// TIA Portal project "1215C_BREAKOUT_BOARD" (V19)

(* hardware
DEVICE "S7-1200 station_1"  S7-1200 Station
   slot 0: "Rack_0"  S7-1200 Rack  Rack  V1.0
   slot 1: "BREAKOUT_BOARD_PLC"  CPU 1215C DC/DC/DC  6ES7 215-1AG40-0XB0  V4.6
DEVICE "BREAKOUT_BOARD_HMI"  KTP400 Basic PN
   slot 0: "BREAKOUT_BOARD_HMI"  KTP400 Basic PN  6AV2 123-2DB03-0AX0  16.0.0.0
   slot 1: "HMI_RT_1"  KTP400 Basic PN  6AV2 123-2DB03-0AX0  16.0.0.0
   slot 5: "BREAKOUT_BOARD_HMI.IE_CP_1"  PROFINET Interface  16.0.0.0
      slot 1: "PROFINET Interface"  PROFINET Interface
         slot 1: "Port_1"  Port
*)

// ===== PLC "BREAKOUT_BOARD_PLC"  CPU 1215C DC/DC/DC =====

VAR_GLOBAL   // PLC tag table "PLC_Outputs"
   "DQ0.0" AT %Q0.0 : Bool;   // Digital Output
   "DQ0.1" AT %Q0.1 : Bool;   // Digital Output
   "DQ0.2" AT %Q0.2 : Bool;   // Digital Output
   "DQ0.3" AT %Q0.3 : Bool;   // Digital Output
   "DQ0.4" AT %Q0.4 : Bool;   // Digital Output
   "DQ0.5" AT %Q0.5 : Bool;   // Digital Output
   "DQ0.6" AT %Q0.6 : Bool;   // Digital Output
   "DQ0.7" AT %Q0.7 : Bool;   // Digital Output
   "DQ1.0" AT %Q1.0 : Bool;   // Digital Output
   "DQ1.1" AT %Q1.1 : Bool;   // Digital Output
   "AQ0.0" AT %QW64 : Word;   // Analog Output
   "AQ0.1" AT %QW66 : Word;   // Analog Output
END_VAR

VAR_GLOBAL   // PLC tag table "PLC_Inputs"
   "DI0.0" AT %I0.0 : Bool;   // Digital Input
   "DI0.1" AT %I0.1 : Bool;   // Digital Input
   "DI0.2" AT %I0.2 : Bool;   // Digital Input
   "DI0.3" AT %I0.3 : Bool;   // Digital Input
   "DI0.4" AT %I0.4 : Bool;   // Digital Input
   "DI0.5" AT %I0.5 : Bool;   // Digital Input
   "DI0.6" AT %I0.6 : Bool;   // Digital Input
   "DI0.7" AT %I0.7 : Bool;   // Digital Input
   "DI1.0" AT %I1.0 : Bool;   // Digital Input
   "DI1.1" AT %I1.1 : Bool;   // Digital Input
   "DI1.2" AT %I1.2 : Bool;   // Digital Input
   "DI1.3" AT %I1.3 : Bool;   // Digital Input
   "DI1.4" AT %I1.4 : Bool;   // Digital Input
   "DI1.5" AT %I1.5 : Bool;   // Digital Input
   "AI0.0" AT %IW64 : Word;   // Analog Input
   "AI0.1" AT %IW66 : Word;   // Analog Input
END_VAR

VAR_GLOBAL   // PLC tag table "System_Tags"
   "Clock_Byte" AT %MB0 : Byte;
   "Clock_10Hz" AT %M0.0 : Bool;
   "Clock_5Hz" AT %M0.1 : Bool;
   "Clock_2.5Hz" AT %M0.2 : Bool;
   "Clock_2Hz" AT %M0.3 : Bool;
   "Clock_1.25Hz" AT %M0.4 : Bool;
   "Clock_1Hz" AT %M0.5 : Bool;
   "Clock_0.625Hz" AT %M0.6 : Bool;
   "Clock_0.5Hz" AT %M0.7 : Bool;
   "System_Byte" AT %MB1 : Byte;
   "FirstScan" AT %M1.0 : Bool;
   "DiagStatusUpdate" AT %M1.1 : Bool;
   "AlwaysTRUE" AT %M1.2 : Bool;
   "AlwaysFALSE" AT %M1.3 : Bool;
END_VAR

VAR_GLOBAL   // PLC tag table "Trigger_Tags"
   "xAQ_Trig" AT %M2.0 : Bool;
   "xTrig2" AT %M2.1 : Bool;
   "xTrig3" AT %M2.2 : Bool;
   "xTrig4" AT %M2.3 : Bool;
   "xTrig5" AT %M2.4 : Bool;
END_VAR

// folder: WS01_TVET_Workstation/00-I/O_Mapping

DATA_BLOCK "DB001-PLC_I/O"   // DB1
{ S7_Optimized_Access := 'TRUE' }
VERSION : 0.1
   VAR
      Inputs : Struct   // PLC Inputs Structure
         "xDI0.0" : Bool;
         "xDI0.1" : Bool;
         "xDI0.2" : Bool;
         "xDI0.3" : Bool;
         "xDI0.4" : Bool;
         "xDI0.5" : Bool;
         "xDI0.6" : Bool;
         "xDI0.7" : Bool;
         "xDI1.0" : Bool;
         "xDI1.1" : Bool;
         "xDI1.2" : Bool;
         "xDI1.3" : Bool;
         "xDI1.4" : Bool;
         "xDI1.5" : Bool;
         "rAI0.0_Scaled" : Real;   // 0 to 24648 = 0 to 10 V
         "rAI0.1_Scaled" : Real;   // 0 to 24648 = 0 to 10 V
      END_STRUCT;
      Outputs : Struct   // PLC Outputs Structure
         "xDQ0.0" : Bool;
         "xDQ0.1" : Bool;
         "xDQ0.2" : Bool;
         "xDQ0.3" : Bool;
         "xDQ0.4" : Bool;
         "xDQ0.5" : Bool;
         "xDQ0.6" : Bool;
         "xDQ0.7" : Bool;
         "xDQ1.0" : Bool;
         "xDQ1.1" : Bool;
         "iAQ0.0_RAW" : Int := 0;
         "rAQ0.0_Scaled" : Real;   // 0 to 24648 = 0 to 20 mA
         "iAQ0.1_RAW" : Int := 0;
         "rAQ0.1_Scaled" : Real;   // 0 to 24648 = 0 to 20 mA
      END_STRUCT;
   END_VAR
BEGIN
END_DATA_BLOCK

// folder: WS01_TVET_Workstation/01-Date_Time

DATA_BLOCK "DB002-DateTime"   // DB2
{ S7_Optimized_Access := 'TRUE' }
VERSION : 0.1
   VAR
      RD_LOC_T_Ret : Int := 0;   // Return value for Read Local Time Block
      LOCAL_DTL : DTL := DTL#1970-01-01-00:00:00;   // RAW DTL
      "Date" : Date := D#1990-01-01;   // RAW Date
      "Time" : Time_Of_Day := TOD#00:00:00;   // RAW Time
      DTLtoString_Ret : String;   // Return value for DTL to String Block
      sCustomDate_YY : String := '';   // Custom year
      sCustomDate_MM : String := '';   // Custom month
      sCustomDate_DD : String := '';   // Custom Day
      sCustomTime_HH : String := '';   // Custom hour
      sCustomTime_MM : String := '';   // Custom minute
      sCustomDate_DDMMYY : String := '';   // Custom date format
      sCustomTime_HHMM : String := '';   // Custom time format
   END_VAR
BEGIN
END_DATA_BLOCK

// folder: (top level)

ORGANIZATION_BLOCK "Main"   // OB1, LAD, ProgramCycle
TITLE = "Main Program Sweep (Cycle)"
{ S7_Optimized_Access := 'TRUE' }
VERSION : 0.1
   VAR_INPUT
      Initial_Call : Bool;   // Initial call of this OB
      Remanence : Bool;   // =True, if remanent data are available
   END_VAR
BEGIN

REGION Network 1 (SCL): ================= PROGRAM_INFORMATION =================
   (*
   ==================================================================
   ********************* PLC I/O BREAKOUT BOARD *********************
   ==================================================================

   TVET Workstation WS01:
   1215C DC/DC/DC - 6ES7215-1AG40-0XB0
   - IP:       192.168.0.175/24

   KTP400 HMI - 6AV2123-2DB03-0AX0
   - IP:       192.168.0.176/24

   =======================================================================

   The program has 2 main sections - I/O Handler & I/O Testing Logic.

   I/O Handler FC:
   We are directly interacting with the PLC's I/O and DB tags, therefore
   a FC is used for the I/O mapping logic.
   - maps the physical inputs & outputs to corresponding tags in DB001,
   - handles scaling of the analog I/O,
   - ensures that physical I/O is only used once in the code.

   I/O Testing Logic FB:
   - Digital inputs can be switched ON/OFF via the HMI or via the physical
     input actuator switches.
   - Digital output states are displayed on the HMI.
   - Analog inputs are controlled via the connected potentiometers.
   - Analog outputs are diplayed on the HMI as a bar graph.

   Additional Notes:
   PLC Tags grouped according to their use/function.

   =======================================================================

   Analog Input Technical data:
   - Number of inputs: 2
   - Type: Voltage (single-ended)
   - Full-scale range: 0 to 10 V
   - Full-scale range (data word): 0 to 27648
   - Overshoot range: 10.001 to 11.759 V
   - Overshoot range (data word): 27649 to 32511
   - Overflow range: 11.760 to 11.852 V
   - Overflow range (data word): 32512 to 32767
   - Resolution: 10 bits
   - Maximum withstand voltage: 35 V DC
   - Smoothing: None, Weak, Medium, or Strong
   - Noise rejection: 10, 50, or 60 Hz
   - Impedance: ≥100 KΩ
   - Isolation (field side to logic): None
   - Accuracy (25 °C / -20 to 60 °C): 3.0% / 3.5% of full-scale
   - Cable length (meters): 100 m, shielded twisted pair
   - Rated range: 0     = 0 V
                  34    = 12 mV
                  20736 = 7.5 V
                  27648 = 10 V

   =======================================================================

   Analog Output Technical data:
   - Number of outputs: 2
   - Type: Current
   - Full-scale range: 0 to 20 mA
   - Full-scale range (data word): 0 to 27648
   - Overshoot range: 20.01 to 23.52 mA
   - Overshoot range (data word): 27649 to 32511
   - Overflow range data word: 32512 to 32767
   - Resolution: 10 bits
   - Output drive impedance: ≤500 Ω max
   - Isolation (field side to logic): None
   - Accuracy (25 °C / -20 to 60 °C): 3.0% / 3.5% of full-scale
   - Settling time: 2 ms
   - Cable length (meters): 100 m, shielded twisted pair
   - Rated range: 0     = 0 mA
                  34    = 0.0247 mA
                  20736 = 15 mA
                  27648 = 20 mA

   =======================================================================
   *)
END_REGION

REGION Network 2: ================= LOCAL_DATE/TIME =================
   // > Call the Date/Time Handler Function
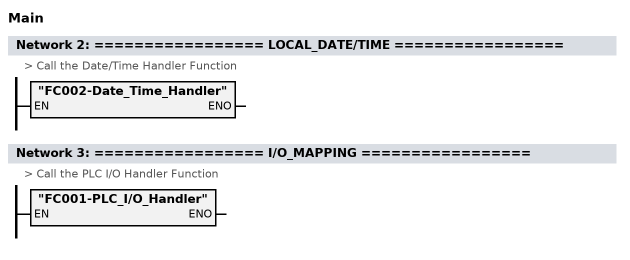
   RUNG wire#powerrail
      "FC002-Date_Time_Handler"()
   END_RUNG
   // the same network as SCL:
   "FC002-Date_Time_Handler"();
END_REGION

REGION Network 3: ================= I/O_MAPPING =================
   // > Call the PLC I/O Handler Function
   RUNG wire#powerrail
      "FC001-PLC_I/O_Handler"()
   END_RUNG
   // the same network as SCL:
   "FC001-PLC_I/O_Handler"();
END_REGION
END_ORGANIZATION_BLOCK

// folder: WS01_TVET_Workstation/00-I/O_Mapping

FUNCTION "FC001-PLC_I/O_Handler" : Void   // FC1, LAD
{ S7_Optimized_Access := 'TRUE' }
VERSION : 0.1
   VAR_TEMP
      "rAI0.0_Temp" : Real;
      "rAI0.1_Temp" : Real;
      "rAQ0.0_Temp" : Real;
      "rAQ0.1_Temp" : Real;
   END_VAR
   VAR_TEMP   // added for the SCL form of the ladder/FBD networks
      _w1 : Bool;
   END_VAR
BEGIN

REGION Network 1: ================= DIGITAL_INPUTS =================
END_REGION

REGION Network 2: BANK_0
   // > DI0.0 - DI0.7
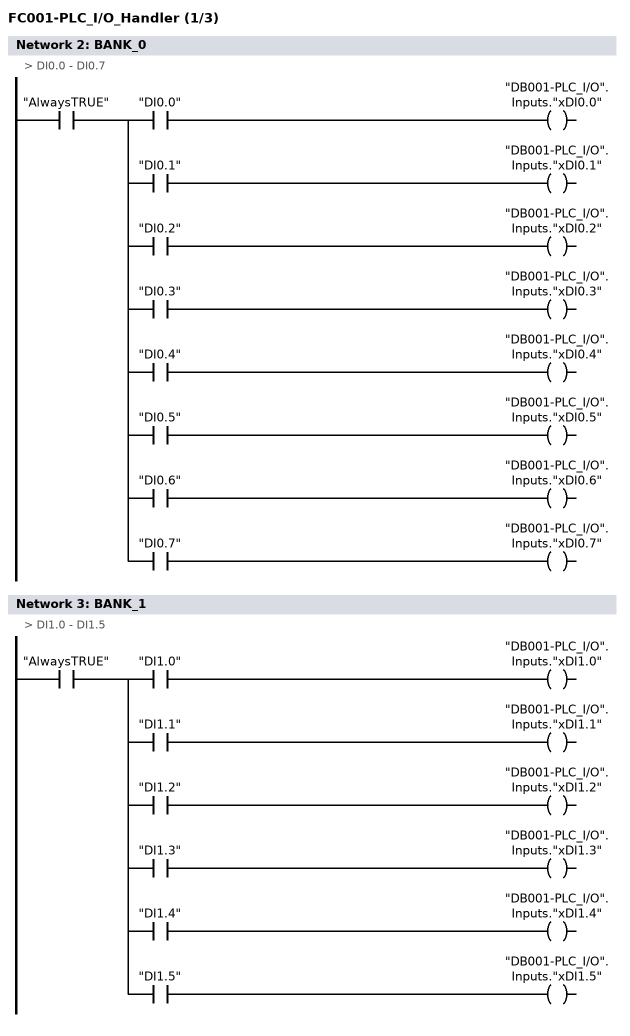
   RUNG wire#powerrail
      Contact( "AlwaysTRUE" )
      wire#w1
      Contact( "DI0.0" )
      Coil( "DB001-PLC_I/O".Inputs."xDI0.0" )
   END_RUNG
   RUNG wire#w1
      Contact( "DI0.1" )
      Coil( "DB001-PLC_I/O".Inputs."xDI0.1" )
   END_RUNG
   RUNG wire#w1
      Contact( "DI0.2" )
      Coil( "DB001-PLC_I/O".Inputs."xDI0.2" )
   END_RUNG
   RUNG wire#w1
      Contact( "DI0.3" )
      Coil( "DB001-PLC_I/O".Inputs."xDI0.3" )
   END_RUNG
   RUNG wire#w1
      Contact( "DI0.4" )
      Coil( "DB001-PLC_I/O".Inputs."xDI0.4" )
   END_RUNG
   RUNG wire#w1
      Contact( "DI0.5" )
      Coil( "DB001-PLC_I/O".Inputs."xDI0.5" )
   END_RUNG
   RUNG wire#w1
      Contact( "DI0.6" )
      Coil( "DB001-PLC_I/O".Inputs."xDI0.6" )
   END_RUNG
   RUNG wire#w1
      Contact( "DI0.7" )
      Coil( "DB001-PLC_I/O".Inputs."xDI0.7" )
   END_RUNG
   // the same network as SCL:
   "DB001-PLC_I/O".Inputs."xDI0.0" := "AlwaysTRUE" AND "DI0.0";
   "DB001-PLC_I/O".Inputs."xDI0.1" := "AlwaysTRUE" AND "DI0.1";
   "DB001-PLC_I/O".Inputs."xDI0.2" := "AlwaysTRUE" AND "DI0.2";
   "DB001-PLC_I/O".Inputs."xDI0.3" := "AlwaysTRUE" AND "DI0.3";
   "DB001-PLC_I/O".Inputs."xDI0.4" := "AlwaysTRUE" AND "DI0.4";
   "DB001-PLC_I/O".Inputs."xDI0.5" := "AlwaysTRUE" AND "DI0.5";
   "DB001-PLC_I/O".Inputs."xDI0.6" := "AlwaysTRUE" AND "DI0.6";
   "DB001-PLC_I/O".Inputs."xDI0.7" := "AlwaysTRUE" AND "DI0.7";
END_REGION

REGION Network 3: BANK_1
   // > DI1.0 - DI1.5
   RUNG wire#powerrail
      Contact( "AlwaysTRUE" )
      wire#w1
      Contact( "DI1.0" )
      Coil( "DB001-PLC_I/O".Inputs."xDI1.0" )
   END_RUNG
   RUNG wire#w1
      Contact( "DI1.1" )
      Coil( "DB001-PLC_I/O".Inputs."xDI1.1" )
   END_RUNG
   RUNG wire#w1
      Contact( "DI1.2" )
      Coil( "DB001-PLC_I/O".Inputs."xDI1.2" )
   END_RUNG
   RUNG wire#w1
      Contact( "DI1.3" )
      Coil( "DB001-PLC_I/O".Inputs."xDI1.3" )
   END_RUNG
   RUNG wire#w1
      Contact( "DI1.4" )
      Coil( "DB001-PLC_I/O".Inputs."xDI1.4" )
   END_RUNG
   RUNG wire#w1
      Contact( "DI1.5" )
      Coil( "DB001-PLC_I/O".Inputs."xDI1.5" )
   END_RUNG
   // the same network as SCL:
   "DB001-PLC_I/O".Inputs."xDI1.0" := "AlwaysTRUE" AND "DI1.0";
   "DB001-PLC_I/O".Inputs."xDI1.1" := "AlwaysTRUE" AND "DI1.1";
   "DB001-PLC_I/O".Inputs."xDI1.2" := "AlwaysTRUE" AND "DI1.2";
   "DB001-PLC_I/O".Inputs."xDI1.3" := "AlwaysTRUE" AND "DI1.3";
   "DB001-PLC_I/O".Inputs."xDI1.4" := "AlwaysTRUE" AND "DI1.4";
   "DB001-PLC_I/O".Inputs."xDI1.5" := "AlwaysTRUE" AND "DI1.5";
END_REGION

REGION Network 4: ================= DIGITAL_OUTPUTS =================
END_REGION

REGION Network 5: BANK_0
   // > DQ0.0 - DQ0.7
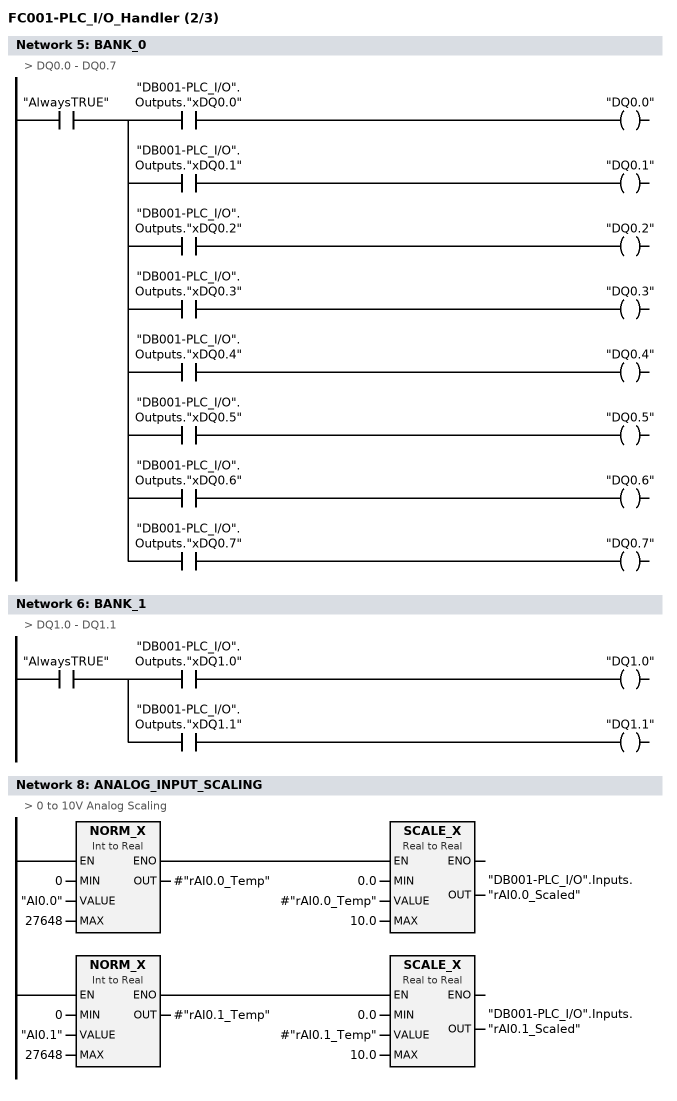
   RUNG wire#powerrail
      Contact( "AlwaysTRUE" )
      wire#w1
      Contact( "DB001-PLC_I/O".Outputs."xDQ0.0" )
      Coil( "DQ0.0" )
   END_RUNG
   RUNG wire#w1
      Contact( "DB001-PLC_I/O".Outputs."xDQ0.1" )
      Coil( "DQ0.1" )
   END_RUNG
   RUNG wire#w1
      Contact( "DB001-PLC_I/O".Outputs."xDQ0.2" )
      Coil( "DQ0.2" )
   END_RUNG
   RUNG wire#w1
      Contact( "DB001-PLC_I/O".Outputs."xDQ0.3" )
      Coil( "DQ0.3" )
   END_RUNG
   RUNG wire#w1
      Contact( "DB001-PLC_I/O".Outputs."xDQ0.4" )
      Coil( "DQ0.4" )
   END_RUNG
   RUNG wire#w1
      Contact( "DB001-PLC_I/O".Outputs."xDQ0.5" )
      Coil( "DQ0.5" )
   END_RUNG
   RUNG wire#w1
      Contact( "DB001-PLC_I/O".Outputs."xDQ0.6" )
      Coil( "DQ0.6" )
   END_RUNG
   RUNG wire#w1
      Contact( "DB001-PLC_I/O".Outputs."xDQ0.7" )
      Coil( "DQ0.7" )
   END_RUNG
   // the same network as SCL:
   "DQ0.0" := "AlwaysTRUE" AND "DB001-PLC_I/O".Outputs."xDQ0.0";
   "DQ0.1" := "AlwaysTRUE" AND "DB001-PLC_I/O".Outputs."xDQ0.1";
   "DQ0.2" := "AlwaysTRUE" AND "DB001-PLC_I/O".Outputs."xDQ0.2";
   "DQ0.3" := "AlwaysTRUE" AND "DB001-PLC_I/O".Outputs."xDQ0.3";
   "DQ0.4" := "AlwaysTRUE" AND "DB001-PLC_I/O".Outputs."xDQ0.4";
   "DQ0.5" := "AlwaysTRUE" AND "DB001-PLC_I/O".Outputs."xDQ0.5";
   "DQ0.6" := "AlwaysTRUE" AND "DB001-PLC_I/O".Outputs."xDQ0.6";
   "DQ0.7" := "AlwaysTRUE" AND "DB001-PLC_I/O".Outputs."xDQ0.7";
END_REGION

REGION Network 6: BANK_1
   // > DQ1.0 - DQ1.1
   RUNG wire#powerrail
      Contact( "AlwaysTRUE" )
      wire#w1
      Contact( "DB001-PLC_I/O".Outputs."xDQ1.0" )
      Coil( "DQ1.0" )
   END_RUNG
   RUNG wire#w1
      Contact( "DB001-PLC_I/O".Outputs."xDQ1.1" )
      Coil( "DQ1.1" )
   END_RUNG
   // the same network as SCL:
   "DQ1.0" := "AlwaysTRUE" AND "DB001-PLC_I/O".Outputs."xDQ1.0";
   "DQ1.1" := "AlwaysTRUE" AND "DB001-PLC_I/O".Outputs."xDQ1.1";
END_REGION

REGION Network 7: ================= ANALOG_PROCESSING =================
END_REGION

REGION Network 8: ANALOG_INPUT_SCALING
   // > 0 to 10V Analog Scaling
   RUNG wire#powerrail
      { S7_Templates := "[SrcType := Int, DestType := Real]" } Normalize(min := 0, value := "AI0.0", max := 27648, out => #"rAI0.0_Temp")
      { S7_Templates := "[SrcType := Real, DestType := Real]" } Scale(min := 0.0, value := #"rAI0.0_Temp", max := 10.0, out => "DB001-PLC_I/O".Inputs."rAI0.0_Scaled")
   END_RUNG
   RUNG wire#powerrail
      { S7_Templates := "[SrcType := Int, DestType := Real]" } Normalize(min := 0, value := "AI0.1", max := 27648, out => #"rAI0.1_Temp")
      { S7_Templates := "[SrcType := Real, DestType := Real]" } Scale(min := 0.0, value := #"rAI0.1_Temp", max := 10.0, out => "DB001-PLC_I/O".Inputs."rAI0.1_Scaled")
   END_RUNG
   // the same network as SCL:
   #"rAI0.0_Temp" := NORM_X(MIN := 0, VALUE := "AI0.0", MAX := 27648);
   "DB001-PLC_I/O".Inputs."rAI0.0_Scaled" := SCALE_X(MIN := 0.0, VALUE := #"rAI0.0_Temp", MAX := 10.0);
   #"rAI0.1_Temp" := NORM_X(MIN := 0, VALUE := "AI0.1", MAX := 27648);
   "DB001-PLC_I/O".Inputs."rAI0.1_Scaled" := SCALE_X(MIN := 0.0, VALUE := #"rAI0.1_Temp", MAX := 10.0);
END_REGION

REGION Network 9: ANALOG_OUTPUT_MANIPULATION
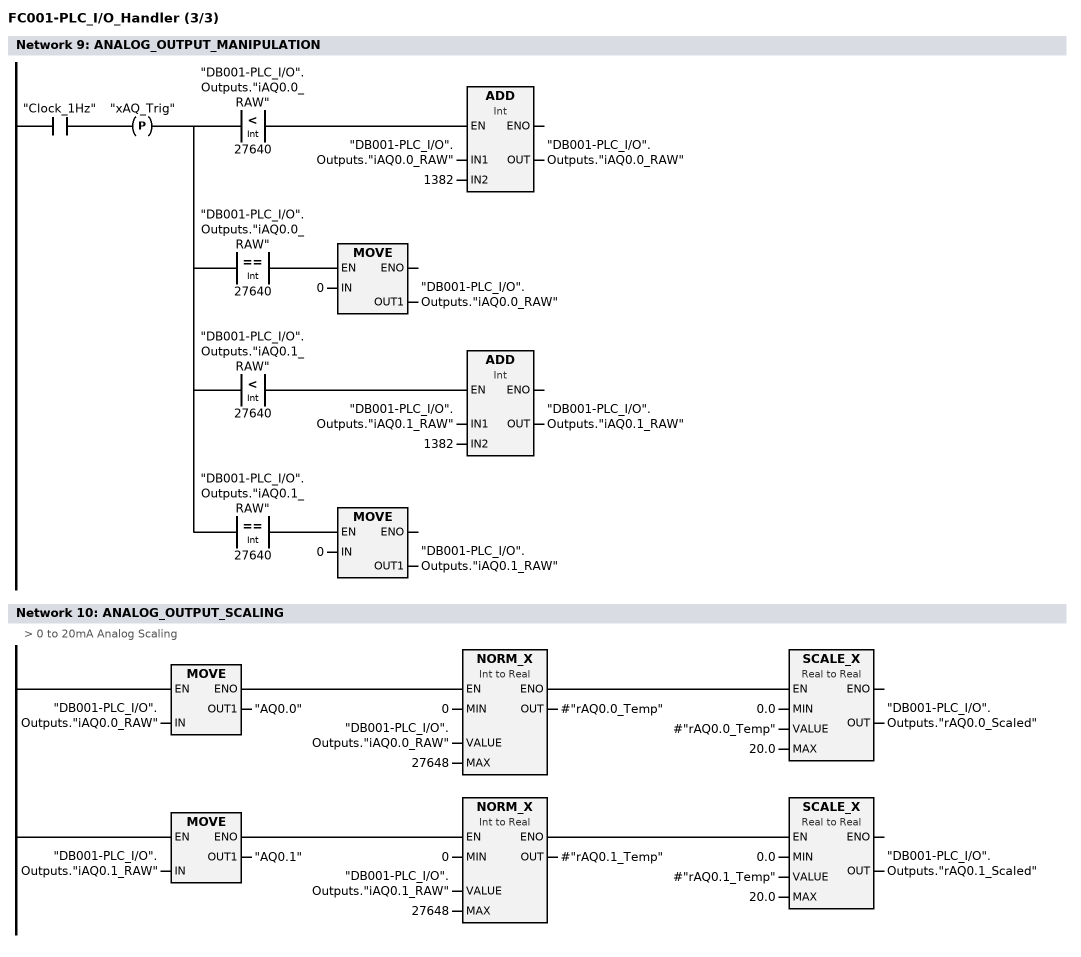
   RUNG wire#powerrail
      Contact( "Clock_1Hz" )
      P_Trig( "xAQ_Trig" )
      wire#w1
      { S7_Templates := "SrcType := Int" } LT_Contact(in1 := "DB001-PLC_I/O".Outputs."iAQ0.0_RAW", in2 := 27640)
      { S7_Templates := "SrcType := Int" } Add(in1 := "DB001-PLC_I/O".Outputs."iAQ0.0_RAW", in2 := 1382, out => "DB001-PLC_I/O".Outputs."iAQ0.0_RAW")
   END_RUNG
   RUNG wire#w1
      { S7_Templates := "SrcType := Int" } EQ_Contact(in1 := "DB001-PLC_I/O".Outputs."iAQ0.0_RAW", in2 := 27640)
      Move(in := 0, out1 => "DB001-PLC_I/O".Outputs."iAQ0.0_RAW")
   END_RUNG
   RUNG wire#w1
      { S7_Templates := "SrcType := Int" } LT_Contact(in1 := "DB001-PLC_I/O".Outputs."iAQ0.1_RAW", in2 := 27640)
      { S7_Templates := "SrcType := Int" } Add(in1 := "DB001-PLC_I/O".Outputs."iAQ0.1_RAW", in2 := 1382, out => "DB001-PLC_I/O".Outputs."iAQ0.1_RAW")
   END_RUNG
   RUNG wire#w1
      { S7_Templates := "SrcType := Int" } EQ_Contact(in1 := "DB001-PLC_I/O".Outputs."iAQ0.1_RAW", in2 := 27640)
      Move(in := 0, out1 => "DB001-PLC_I/O".Outputs."iAQ0.1_RAW")
   END_RUNG
   // the same network as SCL:
   #_w1 := "Clock_1Hz" AND NOT "xAQ_Trig";   // rising edge
   "xAQ_Trig" := "Clock_1Hz";
   IF #_w1 AND ("DB001-PLC_I/O".Outputs."iAQ0.0_RAW" < 27640) THEN
       "DB001-PLC_I/O".Outputs."iAQ0.0_RAW" := "DB001-PLC_I/O".Outputs."iAQ0.0_RAW" + 1382;
   END_IF;
   IF #_w1 AND ("DB001-PLC_I/O".Outputs."iAQ0.0_RAW" = 27640) THEN
       "DB001-PLC_I/O".Outputs."iAQ0.0_RAW" := 0;
   END_IF;
   IF #_w1 AND ("DB001-PLC_I/O".Outputs."iAQ0.1_RAW" < 27640) THEN
       "DB001-PLC_I/O".Outputs."iAQ0.1_RAW" := "DB001-PLC_I/O".Outputs."iAQ0.1_RAW" + 1382;
   END_IF;
   IF #_w1 AND ("DB001-PLC_I/O".Outputs."iAQ0.1_RAW" = 27640) THEN
       "DB001-PLC_I/O".Outputs."iAQ0.1_RAW" := 0;
   END_IF;
END_REGION

REGION Network 10: ANALOG_OUTPUT_SCALING
   // > 0 to 20mA Analog Scaling
   RUNG wire#powerrail
      Move(in := "DB001-PLC_I/O".Outputs."iAQ0.0_RAW", out1 => "AQ0.0")
      { S7_Templates := "[SrcType := Int, DestType := Real]" } Normalize(min := 0, value := "DB001-PLC_I/O".Outputs."iAQ0.0_RAW", max := 27648, out => #"rAQ0.0_Temp")
      { S7_Templates := "[SrcType := Real, DestType := Real]" } Scale(min := 0.0, value := #"rAQ0.0_Temp", max := 20.0, out => "DB001-PLC_I/O".Outputs."rAQ0.0_Scaled")
   END_RUNG
   RUNG wire#powerrail
      Move(in := "DB001-PLC_I/O".Outputs."iAQ0.1_RAW", out1 => "AQ0.1")
      { S7_Templates := "[SrcType := Int, DestType := Real]" } Normalize(min := 0, value := "DB001-PLC_I/O".Outputs."iAQ0.1_RAW", max := 27648, out => #"rAQ0.1_Temp")
      { S7_Templates := "[SrcType := Real, DestType := Real]" } Scale(min := 0.0, value := #"rAQ0.1_Temp", max := 20.0, out => "DB001-PLC_I/O".Outputs."rAQ0.1_Scaled")
   END_RUNG
   // the same network as SCL:
   "AQ0.0" := "DB001-PLC_I/O".Outputs."iAQ0.0_RAW";
   #"rAQ0.0_Temp" := NORM_X(MIN := 0, VALUE := "DB001-PLC_I/O".Outputs."iAQ0.0_RAW", MAX := 27648);
   "DB001-PLC_I/O".Outputs."rAQ0.0_Scaled" := SCALE_X(MIN := 0.0, VALUE := #"rAQ0.0_Temp", MAX := 20.0);
   "AQ0.1" := "DB001-PLC_I/O".Outputs."iAQ0.1_RAW";
   #"rAQ0.1_Temp" := NORM_X(MIN := 0, VALUE := "DB001-PLC_I/O".Outputs."iAQ0.1_RAW", MAX := 27648);
   "DB001-PLC_I/O".Outputs."rAQ0.1_Scaled" := SCALE_X(MIN := 0.0, VALUE := #"rAQ0.1_Temp", MAX := 20.0);
END_REGION
END_FUNCTION

// folder: WS01_TVET_Workstation/01-Date_Time

FUNCTION "FC002-Date_Time_Handler" : Void   // FC2, LAD
{ S7_Optimized_Access := 'TRUE' }
VERSION : 0.1
   VAR_TEMP   // added for the SCL form of the ladder/FBD networks
      _w1 : Bool;
   END_VAR
BEGIN

REGION Network 1: Read Local Date/Time
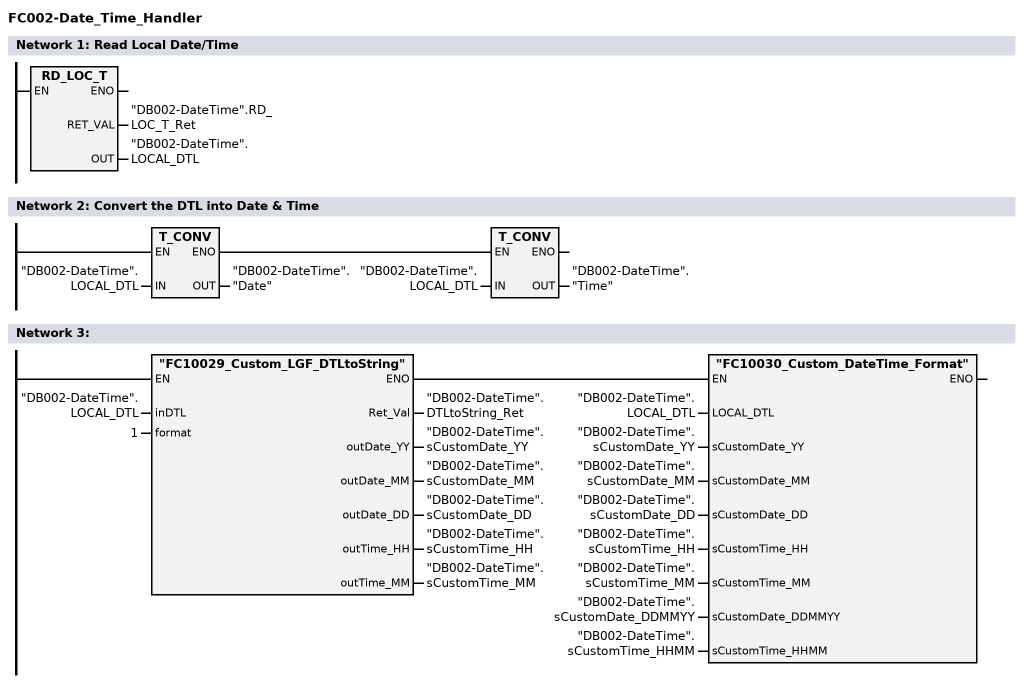
   "DB002-DateTime".RD_LOC_T_Ret := RD_LOC_T(OUT => "DB002-DateTime".LOCAL_DTL);
END_REGION

REGION Network 2: Convert the DTL into Date & Time
   // ENO of a box is taken as its EN; it also drops when the box reports an error
   "DB002-DateTime"."Date" := T_CONV(IN := "DB002-DateTime".LOCAL_DTL);
   "DB002-DateTime"."Time" := T_CONV(IN := "DB002-DateTime".LOCAL_DTL);
END_REGION
